// TIA Portal project "MANF386_lab3_OpPanel" (V16)

(* hardware
DEVICE "S71500/ET200MP station_1"  S7-1500 station
   slot 0: "Rail_0"  Rack  6ES7 590-1***0-0AA0
   slot 1: "PLC_1"  CPU 1512C-1 PN  6ES7 512-1CK00-0AB0  V2.8
      slot 3: "CPU display_1"  6ES7591-1AA00-0AA0
      slot 32768: "PROFINET interface_1"  X1
         slot 32769: "Port_1"  X1 P1
         slot 32770: "Port_2"  X1 P2
      slot 34817: "Virtual CP interface port_1"  Virtual CP interface port  Virtual CP interface port
*)

// ===== PLC "PLC_1"  CPU 1512C-1 PN =====

VAR_GLOBAL   // PLC tag table "Default tag table"
   "start" AT %I11.0 : Bool;
   "stop" AT %I11.1 : Bool;
   "key" AT %I11.2 : Bool;
   "reset" AT %I11.3 : Bool;
   "start_LED" AT %Q5.0 : Bool;
   "reset_LED" AT %Q5.1 : Bool;
   "conv_fwd" AT %Q4.0 : Bool;
   "System_Byte" AT %MB1 : Byte;
   "FirstScan" AT %M1.0 : Bool;
   "DiagStatusUpdate" AT %M1.1 : Bool;
   "AlwaysTRUE" AT %M1.2 : Bool;
   "AlwaysFALSE" AT %M1.3 : Bool;
   "Clock_Byte" AT %MB0 : Byte;
   "Clock_10Hz" AT %M0.0 : Bool;
   "Clock_5Hz" AT %M0.1 : Bool;
   "Clock_2.5Hz" AT %M0.2 : Bool;
   "Clock_2Hz" AT %M0.3 : Bool;
   "Clock_1.25Hz" AT %M0.4 : Bool;
   "Clock_1Hz" AT %M0.5 : Bool;
   "Clock_0.625Hz" AT %M0.6 : Bool;
   "Clock_0.5Hz" AT %M0.7 : Bool;
   "conv_bwd" AT %Q4.1 : Bool;
END_VAR

DATA_BLOCK "controlPanel_DB"   // DB1
{ S7_Optimized_Access := 'TRUE' }
VERSION : 0.1
// stored: InstanceOfName controlPanel
"controlPanel"
BEGIN
END_DATA_BLOCK

FUNCTION_BLOCK "controlPanel"   // FB1, LAD
{ S7_Optimized_Access := 'TRUE' }
VERSION : 0.1
   VAR_INPUT
      start : Bool;
      stop : Bool;
      reset : Bool;
      key : Bool;
   END_VAR
   VAR_OUTPUT
      start_LED : Bool;
      reset_LED : Bool;
      conv_fwd : Bool;
   END_VAR
   VAR
      state1 : Bool;
      state2 : Bool;
      edge1 : Bool;
      edge2 : Bool;
      state4 : Bool;
      state3 : Bool;
   END_VAR
   VAR_TEMP
      tr1_2 : Bool;
      key_change : Bool;
      tr2_1 : Bool;
      tr2_4 : Bool;
      tr2_3 : Bool;
      tr4_1 : Bool;
      tr3_2 : Bool;
      tr3_1 : Bool;
   END_VAR
   VAR_TEMP   // added for the SCL form of the ladder/FBD networks
      _w1 : Bool;
      _w2 : Bool;
   END_VAR
BEGIN

REGION Network 1: key change
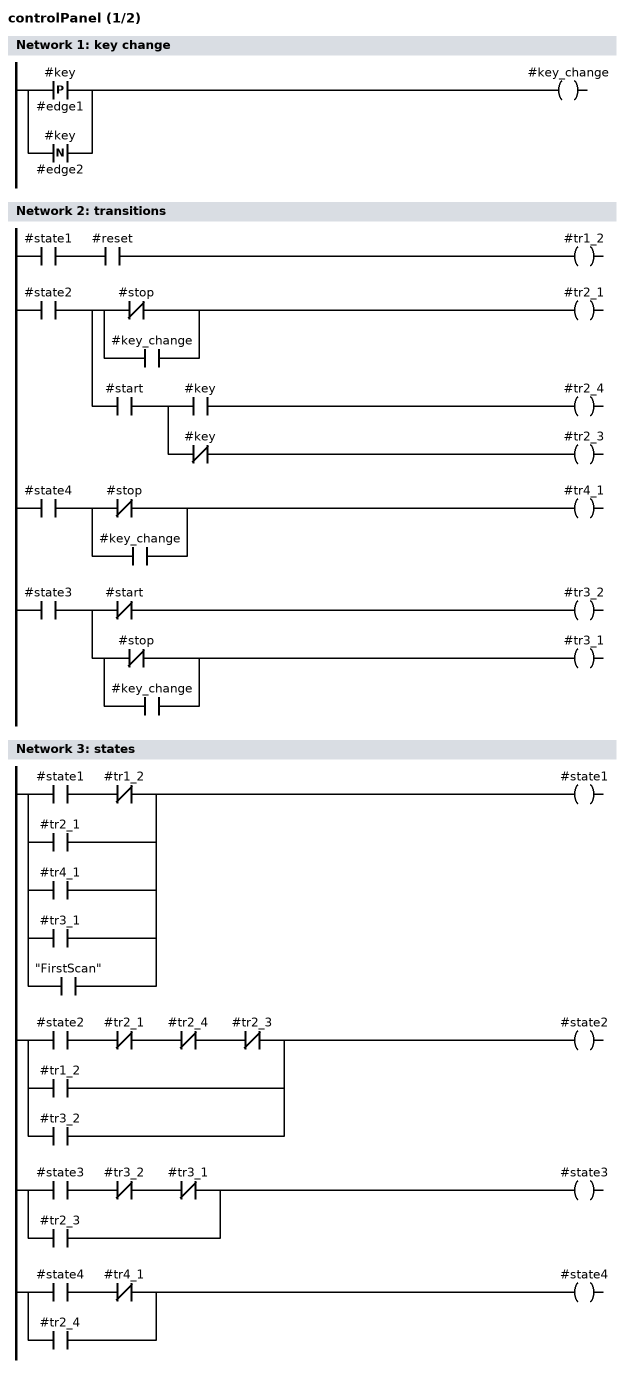
   RUNG wire#powerrail
      P_Contact(operand := #key, bit := #edge1)
      wire#w1
      Coil( #key_change )
   END_RUNG
   RUNG wire#powerrail
      N_Contact(operand := #key, bit := #edge2)
   END_RUNG wire#w1
   // the same network as SCL:
   #_w1 := #key AND NOT #edge1;   // rising edge of #key
   #edge1 := #key;
   #_w2 := NOT #key AND #edge2;   // falling edge of #key
   #edge2 := #key;
   #key_change := #_w1 OR #_w2;
END_REGION

REGION Network 2: transitions
   RUNG wire#powerrail
      Contact( #state1 )
      Contact( #reset )
      Coil( #tr1_2 )
   END_RUNG
   RUNG wire#powerrail
      Contact( #state2 )
      wire#w1
      I_Contact( #stop )
      wire#w2
      Coil( #tr2_1 )
   END_RUNG
   RUNG wire#w1
      Contact( #key_change )
   END_RUNG wire#w2
   RUNG wire#w1
      Contact( #start )
      wire#w3
      Contact( #key )
      Coil( #tr2_4 )
   END_RUNG
   RUNG wire#w3
      I_Contact( #key )
      Coil( #tr2_3 )
   END_RUNG
   RUNG wire#powerrail
      Contact( #state4 )
      wire#w4
      I_Contact( #stop )
      wire#w5
      Coil( #tr4_1 )
   END_RUNG
   RUNG wire#w4
      Contact( #key_change )
   END_RUNG wire#w5
   RUNG wire#powerrail
      Contact( #state3 )
      wire#w6
      I_Contact( #start )
      Coil( #tr3_2 )
   END_RUNG
   RUNG wire#w6
      I_Contact( #stop )
      wire#w7
      Coil( #tr3_1 )
   END_RUNG
   RUNG wire#w6
      Contact( #key_change )
   END_RUNG wire#w7
   // the same network as SCL:
   #tr1_2 := #state1 AND #reset;
   #tr2_1 := #state2 AND (NOT #stop OR #key_change);
   #_w1 := #state2 AND #start;
   #tr2_4 := #_w1 AND #key;
   #tr2_3 := #_w1 AND NOT #key;
   #tr4_1 := #state4 AND (NOT #stop OR #key_change);
   #tr3_2 := #state3 AND NOT #start;
   #tr3_1 := #state3 AND (NOT #stop OR #key_change);
END_REGION

REGION Network 3: states
   RUNG wire#powerrail
      Contact( #state1 )
      I_Contact( #tr1_2 )
      wire#w1
      Coil( #state1 )
   END_RUNG
   RUNG wire#powerrail
      Contact( #tr2_1 )
   END_RUNG wire#w1
   RUNG wire#powerrail
      Contact( #tr4_1 )
   END_RUNG wire#w1
   RUNG wire#powerrail
      Contact( #tr3_1 )
   END_RUNG wire#w1
   RUNG wire#powerrail
      Contact( "FirstScan" )
   END_RUNG wire#w1
   RUNG wire#powerrail
      Contact( #state2 )
      I_Contact( #tr2_1 )
      I_Contact( #tr2_4 )
      I_Contact( #tr2_3 )
      wire#w2
      Coil( #state2 )
   END_RUNG
   RUNG wire#powerrail
      Contact( #tr1_2 )
   END_RUNG wire#w2
   RUNG wire#powerrail
      Contact( #tr3_2 )
   END_RUNG wire#w2
   RUNG wire#powerrail
      Contact( #state3 )
      I_Contact( #tr3_2 )
      I_Contact( #tr3_1 )
      wire#w3
      Coil( #state3 )
   END_RUNG
   RUNG wire#powerrail
      Contact( #tr2_3 )
   END_RUNG wire#w3
   RUNG wire#powerrail
      Contact( #state4 )
      I_Contact( #tr4_1 )
      wire#w4
      Coil( #state4 )
   END_RUNG
   RUNG wire#powerrail
      Contact( #tr2_4 )
   END_RUNG wire#w4
   // the same network as SCL:
   #state1 := (#state1 AND NOT #tr1_2) OR #tr2_1 OR #tr4_1 OR #tr3_1 OR "FirstScan";
   #state2 := (#state2 AND NOT #tr2_1 AND NOT #tr2_4 AND NOT #tr2_3) OR #tr1_2 OR #tr3_2;
   #state3 := (#state3 AND NOT #tr3_2 AND NOT #tr3_1) OR #tr2_3;
   #state4 := (#state4 AND NOT #tr4_1) OR #tr2_4;
END_REGION

REGION Network 4: state logic
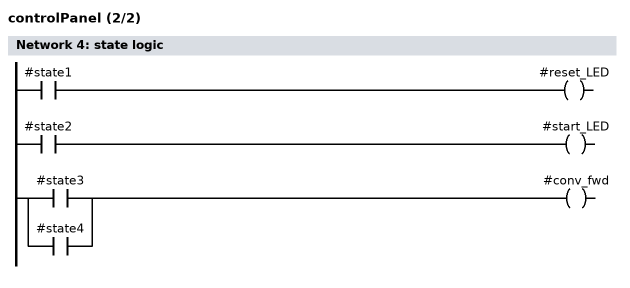
   RUNG wire#powerrail
      Contact( #state1 )
      Coil( #reset_LED )
   END_RUNG
   RUNG wire#powerrail
      Contact( #state2 )
      Coil( #start_LED )
   END_RUNG
   RUNG wire#powerrail
      Contact( #state3 )
      wire#w1
      Coil( #conv_fwd )
   END_RUNG
   RUNG wire#powerrail
      Contact( #state4 )
   END_RUNG wire#w1
   // the same network as SCL:
   #reset_LED := #state1;
   #start_LED := #state2;
   #conv_fwd := #state3 OR #state4;
END_REGION
END_FUNCTION_BLOCK

ORGANIZATION_BLOCK "Main"   // OB1, LAD, ProgramCycle
TITLE = "Main Program Sweep (Cycle)"
{ S7_Optimized_Access := 'TRUE' }
VERSION : 0.1
   VAR_INPUT
      Initial_Call : Bool;   // Initial call of this OB
      Remanence : Bool;   // =True, if remanent data are available
   END_VAR
BEGIN

REGION Network 1
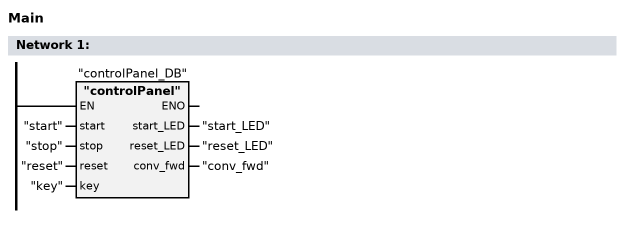
   RUNG wire#powerrail
      "controlPanel_DB"(start := "start", stop := "stop", reset := "reset", key := "key", start_LED => "start_LED", reset_LED => "reset_LED", conv_fwd => "conv_fwd")
   END_RUNG
   // the same network as SCL:
   "controlPanel_DB"(start := "start",   // "controlPanel"
                     stop := "stop",
                     reset := "reset",
                     key := "key",
                     start_LED => "start_LED",
                     reset_LED => "reset_LED",
                     conv_fwd => "conv_fwd");
END_REGION
END_ORGANIZATION_BLOCK